      Appearance <- "VP 45"
   Polygon "Polygon_196" at 843,458 size 11x11
      Appearance <- "VP 45"
   Polygon "Polygon_199" at 630,469 size 11x11
      Appearance <- "VP 33"
   Polygon "Polygon_200" at 631,458 size 11x11
      Appearance <- "VP 33"
   Polygon "Polygon_157" at 417,469 size 11x11
      Appearance <- "VP 21"
   Polygon "Polygon_158" at 418,458 size 11x11
      Appearance <- "VP 21"
   Polygon "Polygon_151" at 205,469 size 11x11
      Appearance <- "VP 16"
   Polygon "Polygon_152" at 206,458 size 11x11
      Appearance <- "VP 16"
   Polygon "Polygon_201" at 83,465 size 11x11
      Appearance <- "VP 1"
   Polygon "Polygon_202" at 94,466 size 11x11
      Appearance <- "VP 1"
   Polygon "Polygon_5" at 83,508 size 11x11
      Appearance <- "VP 2"
   Polygon "Polygon_6" at 94,509 size 11x11
      Appearance <- "VP 2"
   Polygon "Polygon_7" at 83,551 size 11x11
      Appearance <- "VP 3"
   Polygon "Polygon_8" at 94,552 size 11x11
      Appearance <- "VP 3"
   Polygon "Polygon_9" at 83,595 size 11x11
      Appearance <- "VP 4"
   Polygon "Polygon_10" at 94,596 size 11x11
      Appearance <- "VP 4"
   Polygon "Polygon_11" at 124,490 size 11x11
      Appearance <- "VP 5"
   Polygon "Polygon_12" at 135,491 size 11x11
      Appearance <- "VP 5"
   Polygon "Polygon_13" at 158,490 size 11x11
      Appearance <- "VP 7"
   Polygon "Polygon_14" at 169,491 size 11x11
      Appearance <- "VP 7"
   Polygon "Polygon_15" at 124,576 size 11x11
      Appearance <- "VP 6"
   Polygon "Polygon_16" at 135,577 size 11x11
      Appearance <- "VP 6"
   Polygon "Polygon_207" at 158,576 size 11x11
      Appearance <- "VP 8"
   Polygon "Polygon_208" at 169,577 size 11x11
      Appearance <- "VP 8"
   Polygon "Polygon_17" at 295,465 size 11x11
      Appearance <- "VP 9"
   Polygon "Polygon_18" at 306,466 size 11x11
      Appearance <- "VP 9"
   Polygon "Polygon_19" at 295,508 size 11x11
      Appearance <- "VP 10"
   Polygon "Polygon_20" at 306,509 size 11x11
      Appearance <- "VP 10"
   Polygon "Polygon_21" at 295,551 size 11x11
      Appearance <- "VP 11"
   Polygon "Polygon_22" at 306,552 size 11x11
      Appearance <- "VP 11"
   Polygon "Polygon_23" at 295,595 size 11x11
      Appearance <- "VP 12"
   Polygon "Polygon_24" at 306,596 size 11x11
      Appearance <- "VP 12"
   Polygon "Polygon_25" at 336,490 size 11x11
      Appearance <- "VP 17"
   Polygon "Polygon_26" at 347,491 size 11x11
      Appearance <- "VP 17"
   Polygon "Polygon_27" at 370,490 size 11x11
      Appearance <- "VP 18"
   Polygon "Polygon_28" at 381,491 size 11x11
      Appearance <- "VP 18"
   Polygon "Polygon_29" at 336,576 size 11x11
      Appearance <- "VP 19"
   Polygon "Polygon_30" at 347,577 size 11x11
      Appearance <- "VP 19"
   Polygon "Polygon_31" at 370,576 size 11x11
      Appearance <- "VP 20"
   Polygon "Polygon_32" at 381,577 size 11x11
      Appearance <- "VP 20"
   Polygon "Polygon_33" at 507,465 size 11x11
      Appearance <- "VP 24"
   Polygon "Polygon_34" at 518,466 size 11x11
      Appearance <- "VP 24"
   Polygon "Polygon_35" at 507,508 size 11x11
      Appearance <- "VP 25"
   Polygon "Polygon_36" at 518,509 size 11x11
      Appearance <- "VP 25"
   Polygon "Polygon_37" at 507,551 size 11x11
      Appearance <- "VP 26"
   Polygon "Polygon_38" at 518,552 size 11x11
      Appearance <- "VP 26"
   Polygon "Polygon_39" at 507,595 size 11x11
      Appearance <- "VP 27"
   Polygon "Polygon_40" at 518,596 size 11x11
      Appearance <- "VP 27"
   Polygon "Polygon_41" at 548,490 size 11x11
      Appearance <- "VP 29"
   Polygon "Polygon_42" at 559,491 size 11x11
      Appearance <- "VP 29"
   Polygon "Polygon_43" at 582,490 size 11x11
      Appearance <- "VP 30"
   Polygon "Polygon_44" at 593,491 size 11x11
      Appearance <- "VP 30"
   Polygon "Polygon_45" at 548,576 size 11x11
      Appearance <- "VP 31"
   Polygon "Polygon_46" at 559,577 size 11x11
      Appearance <- "VP 31"
   Polygon "Polygon_47" at 582,576 size 11x11
      Appearance <- "VP 32"
   Polygon "Polygon_48" at 593,577 size 11x11
      Appearance <- "VP 32"
   Polygon "Polygon_49" at 719,465 size 11x11
      Appearance <- "VP 36"
   Polygon "Polygon_50" at 730,466 size 11x11
      Appearance <- "VP 36"
   Polygon "Polygon_51" at 719,508 size 11x11
      Appearance <- "VP 37"
   Polygon "Polygon_52" at 730,509 size 11x11
      Appearance <- "VP 37"
   Polygon "Polygon_53" at 719,551 size 11x11
      Appearance <- "VP 38"
   Polygon "Polygon_54" at 730,552 size 11x11
      Appearance <- "VP 38"
   Polygon "Polygon_55" at 719,595 size 11x11
      Appearance <- "VP 39"
   Polygon "Polygon_56" at 730,596 size 11x11
      Appearance <- "VP 39"
   Polygon "Polygon_57" at 760,490 size 11x11
      Appearance <- "VP 41"
   Polygon "Polygon_58" at 771,491 size 11x11
      Appearance <- "VP 41"
   Polygon "Polygon_59" at 794,490 size 11x11
      Appearance <- "VP 42"
   Polygon "Polygon_60" at 805,491 size 11x11
      Appearance <- "VP 42"
   Polygon "Polygon_61" at 760,576 size 11x11
      Appearance <- "VP 43"
   Polygon "Polygon_62" at 771,577 size 11x11
      Appearance <- "VP 43"
   Polygon "Polygon_63" at 794,576 size 11x11
      Appearance <- "VP 44"
   Polygon "Polygon_64" at 805,577 size 11x11
      Appearance <- "VP 44"
   Polygon "Polygon_65" at 931,465 size 11x11
      Appearance <- "VP 48"
   Polygon "Polygon_66" at 942,466 size 11x11
      Appearance <- "VP 48"
   Polygon "Polygon_67" at 931,508 size 11x11
      Appearance <- "VP 49"
   Polygon "Polygon_68" at 942,509 size 11x11
      Appearance <- "VP 49"
   Polygon "Polygon_69" at 931,551 size 11x11
      Appearance <- "VP 50"
   Polygon "Polygon_70" at 942,552 size 11x11
      Appearance <- "VP 50"
   Polygon "Polygon_71" at 931,595 size 11x11
      Appearance <- "VP 51"
   Polygon "Polygon_72" at 942,596 size 11x11
      Appearance <- "VP 51"
   Polygon "Polygon_73" at 972,490 size 11x11
      Appearance <- "VP 53"
   Polygon "Polygon_74" at 983,491 size 11x11
      Appearance <- "VP 53"
   Polygon "Polygon_75" at 1006,490 size 11x11
      Appearance <- "VP 54"
   Polygon "Polygon_76" at 1017,491 size 11x11
      Appearance <- "VP 54"
   Polygon "Polygon_77" at 972,576 size 11x11
      Appearance <- "VP 55"
   Polygon "Polygon_78" at 983,577 size 11x11
      Appearance <- "VP 55"
   Polygon "Polygon_79" at 1006,576 size 11x11
      Appearance <- "VP 56"
   Polygon "Polygon_80" at 1017,577 size 11x11
      Appearance <- "VP 56"
   Polygon "Polygon_81" at 1143,465 size 11x11
      Appearance <- "VP 60"
   Polygon "Polygon_82" at 1154,466 size 11x11
      Appearance <- "VP 60"
   Polygon "Polygon_83" at 1143,508 size 11x11
      Appearance <- "VP 61"
   Polygon "Polygon_84" at 1154,509 size 11x11
      Appearance <- "VP 61"
   Polygon "Polygon_85" at 1143,551 size 11x11
      Appearance <- "VP 62"
   Polygon "Polygon_86" at 1154,552 size 11x11
      Appearance <- "VP 62"
   Polygon "Polygon_87" at 1143,595 size 11x11
      Appearance <- "VP 63"
   Polygon "Polygon_88" at 1154,596 size 11x11
      Appearance <- "VP 63"
   Polygon "Polygon_89" at 1184,490 size 11x11
      Appearance <- "VP 65"
   Polygon "Polygon_90" at 1195,491 size 11x11
      Appearance <- "VP 65"
   Polygon "Polygon_91" at 1218,490 size 11x11
      Appearance <- "VP 66"
   Polygon "Polygon_92" at 1229,491 size 11x11
      Appearance <- "VP 66"
   Polygon "Polygon_93" at 1184,576 size 11x11
      Appearance <- "VP 67"
   Polygon "Polygon_94" at 1195,577 size 11x11
      Appearance <- "VP 67"
   Polygon "Polygon_95" at 1218,576 size 11x11
      Appearance <- "VP 68"
   Polygon "Polygon_96" at 1229,577 size 11x11
      Appearance <- "VP 68"
   Polygon "Polygon_97" at 1355,465 size 11x11
      Appearance <- "VP 72"
   Polygon "Polygon_98" at 1366,466 size 11x11
      Appearance <- "VP 72"
   Polygon "Polygon_99" at 1355,508 size 11x11
      Appearance <- "VP 73"
   Polygon "Polygon_100" at 1366,509 size 11x11
      Appearance <- "VP 73"
   Polygon "Polygon_101" at 1355,551 size 11x11
      Appearance <- "VP 74"
   Polygon "Polygon_102" at 1366,552 size 11x11
      Appearance <- "VP 74"
   Polygon "Polygon_103" at 1355,595 size 11x11
      Appearance <- "VP 75"
   Polygon "Polygon_104" at 1366,596 size 11x11
      Appearance <- "VP 75"
   Polygon "Polygon_105" at 1396,490 size 11x11
      Appearance <- "VP 77"
   Polygon "Polygon_106" at 1407,491 size 11x11
      Appearance <- "VP 77"
   Polygon "Polygon_107" at 1430,490 size 11x11
      Appearance <- "VP 78"
   Polygon "Polygon_108" at 1441,491 size 11x11
      Appearance <- "VP 78"
   Polygon "Polygon_109" at 1396,576 size 11x11
      Appearance <- "VP 79"
   Polygon "Polygon_110" at 1407,577 size 11x11
      Appearance <- "VP 79"
   Polygon "Polygon_111" at 1430,576 size 11x11
      Appearance <- "VP 80"
   Polygon "Polygon_112" at 1441,577 size 11x11
      Appearance <- "VP 80"
   Polygon "Polygon_113" at 142,942 size 11x11
      Appearance <- "VP 87"
   Polygon "Polygon_114" at 153,943 size 11x11
      Appearance <- "VP 87"
   Polygon "Polygon_3" at 30,890 size 11x11
      Appearance <- "VP 86"
   Polygon "Polygon_4" at 41,891 size 11x11
      Appearance <- "VP 86"
   Polygon "Polygon_115" at 123,352 size 58x419
      Visibility <- "step_vessel_1_proses"
      Appearance <- "VP 5"
   Line "Line_112" at 124,432 size 57x0
      Visibility <- "step_vessel_1_proses"
   Line "Line_113" at 142,385 size 21x0
      Visibility <- "step_vessel_1_proses"
   Line "Line_114" at 124,680 size 56x0
      Visibility <- "step_vessel_1_proses"
   Polygon "Polygon_116" at 335,352 size 58x419
      Appearance <- "VP 17"
      Visibility <- "step_vessel_2_proses"
   Line "Line_115" at 336,432 size 57x0
      Visibility <- "step_vessel_2_proses"
   Line "Line_116" at 354,385 size 21x0
      Visibility <- "step_vessel_2_proses"
   Line "Line_211" at 336,680 size 56x0
      Visibility <- "step_vessel_2_proses"
   Polygon "Polygon_189" at 547,352 size 58x419
      Appearance <- "VP 29"
      Visibility <- "step_vessel_3_proses"
   Line "Line_212" at 548,432 size 57x0
      Visibility <- "step_vessel_3_proses"
   Line "Line_213" at 566,385 size 21x0
      Visibility <- "step_vessel_3_proses"
   Line "Line_214" at 548,680 size 56x0
      Visibility <- "step_vessel_3_proses"
   Polygon "Polygon_190" at 759,352 size 58x419
      Appearance <- "VP 41"
      Visibility <- "step_vessel_4_proses"
   Line "Line_215" at 760,432 size 57x0
      Visibility <- "step_vessel_4_proses"
   Line "Line_216" at 778,385 size 21x0
      Visibility <- "step_vessel_4_proses"
   Line "Line_217" at 760,680 size 56x0
      Visibility <- "step_vessel_4_proses"
   Polygon "Polygon_203" at 971,352 size 58x419
      Appearance <- "VP 53"
      Visibility <- "step_vessel_5_proses"
   Line "Line_218" at 972,432 size 57x0
      Visibility <- "step_vessel_5_proses"
   Line "Line_219" at 990,385 size 21x0
      Visibility <- "step_vessel_5_proses"
   Line "Line_220" at 972,680 size 56x0
      Visibility <- "step_vessel_5_proses"
   Polygon "Polygon_204" at 1183,352 size 58x419
      Appearance <- "VP 65"
      Visibility <- "step_vessel_6_proses"
   Line "Line_221" at 1184,432 size 57x0
      Visibility <- "step_vessel_6_proses"
   Line "Line_222" at 1202,385 size 21x0
      Visibility <- "step_vessel_6_proses"
   Line "Line_223" at 1184,680 size 56x0
      Visibility <- "step_vessel_6_proses"
   Polygon "Polygon_209" at 1395,352 size 58x419
      Appearance <- "VP 77"
      Visibility <- "step_vessel_7_proses"
   Line "Line_224" at 1396,432 size 57x0
      Visibility <- "step_vessel_7_proses"
   Line "Line_225" at 1414,385 size 21x0
      Visibility <- "step_vessel_7_proses"
   Line "Line_226" at 1396,680 size 56x0
      Visibility <- "step_vessel_7_proses"
   IOField "I/O field_3" at 141,608 size 38x17; FormatPattern 9999999
   TextField "Text field_15" at 177,608 size 25x18; Text 'bar'
   IOField "I/O field_4" at 141,632 size 38x17; FormatPattern 9999999
   TextField "Text field_16" at 177,632 size 23x18; Text 'º C'
   IOField "I/O field_7" at 353,608 size 38x17; FormatPattern 9999999
   TextField "Text field_31" at 389,608 size 25x18; Text 'bar'
   IOField "I/O field_8" at 353,632 size 38x17; FormatPattern 9999999
   TextField "Text field_32" at 389,632 size 23x18; Text 'º C'
   IOField "I/O field_11" at 565,608 size 38x17; FormatPattern 9999999
   TextField "Text field_5" at 601,608 size 25x18; Text 'bar'
   IOField "I/O field_12" at 565,632 size 38x17; FormatPattern 9999999
   TextField "Text field_6" at 601,632 size 23x18; Text 'º C'
   IOField "I/O field_15" at 777,608 size 38x17; FormatPattern 9999999
   TextField "Text field_17" at 813,608 size 25x18; Text 'bar'
   IOField "I/O field_16" at 777,632 size 38x17; FormatPattern 9999999
   TextField "Text field_18" at 813,632 size 23x18; Text 'º C'
   IOField "I/O field_19" at 989,608 size 38x17; FormatPattern 9999999
   TextField "Text field_19" at 1025,608 size 25x18; Text 'bar'
   IOField "I/O field_20" at 989,632 size 38x17; FormatPattern 9999999
   TextField "Text field_20" at 1025,632 size 23x18; Text 'º C'
   IOField "I/O field_23" at 1201,608 size 38x17; FormatPattern 9999999
   TextField "Text field_21" at 1237,608 size 25x18; Text 'bar'
   IOField "I/O field_24" at 1201,632 size 38x17; FormatPattern 9999999
   TextField "Text field_22" at 1237,632 size 23x18; Text 'º C'
   IOField "I/O field_27" at 1413,608 size 38x17; FormatPattern 9999999
   TextField "Text field_23" at 1449,608 size 25x18; Text 'bar'
   IOField "I/O field_28" at 1413,632 size 38x17; FormatPattern 9999999
   TextField "Text field_24" at 1449,632 size 23x18; Text 'º C'
   Line "Line_1" at 109,467 size 0x141
      Appearance <- "step_vessel_1"
      Visibility <- "step_vessel_1_proses"
   Line "Line_3" at 110,496 size 16x0
      Appearance <- "step_vessel_1"
      Visibility <- "step_vessel_1_proses"
   Line "Line_4" at 110,582 size 16x0
      Appearance <- "step_vessel_1"
      Visibility <- "step_vessel_1_proses"
   Line "Line_17" at 321,466 size 0x157
      Appearance <- "step_vessel_2"
      Visibility <- "step_vessel_2_proses"
   Line "Line_18" at 318,496 size 16x0
      Appearance <- "step_vessel_2"
      Visibility <- "step_vessel_2_proses"
   Line "Line_19" at 318,582 size 16x0
      Appearance <- "step_vessel_2"
      Visibility <- "step_vessel_2_proses"
   Group "Tank vessel 1_1" at 123,352 size 58x419
   Group "Group_1" at 109,467 size 17x141
   Group "Group_76" at 180,475 size 118x150
   Group "Group_100" at 318,466 size 16x157
   Group "Tank vessel 2_1" at 335,352 size 58x419
   Group "Group_126" at 392,475 size 118x150
   Group "Group_148" at 605,475 size 118x150
   Group "Group_149" at 817,475 size 118x150
   Group "Group_150" at 1030,475 size 118x150
   Group "Group_151" at 1241,475 size 114x150
   Group "Group_152" at 1453,481 size 80x138
   Group "Group_86" at 739,620 size 12x22
   Group "Group_157" at 745,466 size 21x155
   Group "Group_155" at 533,466 size 17x154
   Group "Group_159" at 954,466 size 20x158
   Group "Group_161" at 1169,466 size 21x156
   Group "Group_163" at 1381,466 size 17x156
   Group "Group_5" at 536,400 size 40x99
   Group "Group_189" at 1172,400 size 40x99
   Polyline "Polyline_8" at 153,793 size 18x84
      Visibility <- "VB 1"
      Appearance <- "step_vessel_1_proses"
   Polyline "Polyline_11" at 365,793 size 18x84
      Visibility <- "VB 2"
      Appearance <- "step_vessel_2_proses"
   Polyline "Polyline_12" at 577,793 size 18x84
      Visibility <- "VB 3"
      Appearance <- "step_vessel_3_proses"
   Polyline "Polyline_14" at 789,793 size 18x84
      Visibility <- "VB 4"
      Appearance <- "step_vessel_4_proses"
   Polyline "Polyline_16" at 1001,793 size 18x84
      Visibility <- "VB 5"
      Appearance <- "step_vessel_5_proses"
   Polyline "Polyline_18" at 1213,793 size 18x84
      Visibility <- "VB 6"
      Appearance <- "step_vessel_6_proses"
   Polyline "Polyline_20" at 1425,793 size 18x84
      Visibility <- "VB 7"
      Appearance <- "step_vessel_7_proses"
   Group "Group_129" at 547,352 size 58x419
   Group "Group_144" at 759,352 size 58x419
   Group "Group_145" at 971,352 size 58x419
   Group "Group_146" at 1183,352 size 58x419
   Group "Group_147" at 1395,352 size 58x419
   Group "Tank vessel 1" at 123,352 size 58x419
   Group "Tank vessel 2" at 335,352 size 58x419
   Group "Group_116" at 547,352 size 58x419
   Group "Group_119" at 759,352 size 58x419
   Group "Group_120" at 971,352 size 58x419
   Group "Group_121" at 1183,352 size 58x419
   Group "Group_122" at 1395,352 size 58x419
   Group "Tank vessel 1_2" at 123,352 size 58x419
   Group "Tank vessel 2_2" at 335,352 size 58x419
   Group "Group_196" at 547,352 size 58x419
   Group "Group_197" at 759,352 size 58x419
   Group "Group_198" at 971,352 size 58x419
   Group "Group_200" at 1395,352 size 58x419
   Group "Group_199" at 1183,352 size 58x419
   Group "Group_127" at 420,640 size 1121x45
   Polygon "Polygon_210" at 123,352 size 58x419
      Visibility <- "step_vessel_1_proses"
      Appearance <- "step_vessel_1_proses"
   Line "Line_110" at 124,432 size 57x0
      Visibility <- "step_vessel_1_proses"
   Line "Line_111" at 142,385 size 21x0
      Visibility <- "step_vessel_1_proses"
   Line "Line_227" at 124,680 size 56x0
      Visibility <- "step_vessel_1_proses"
   Line "Line_228" at 112,400 size 25x11
      Visibility <- "VP 5"
      Appearance <- "step_vessel_1_proses"
   Line "Line_229" at 116,412 size 36x78
      Visibility <- "VP 5"
      Appearance <- "step_vessel_1_proses"
   Line "Line_230" at 152,488 size 0x11
      Visibility <- "VP 5"
      Appearance <- "step_vessel_1_proses"
   Line "Line_232" at 131,595 size 21x144
      Visibility <- "VP 5"
      Appearance <- "step_vessel_1_proses"
   Line "Line_233" at 152,579 size 0x19
      Visibility <- "VP 5"
      Appearance <- "step_vessel_1_proses"
   Line "Line_234" at 128,739 size 25x0
      Visibility <- "VP 5"
      Appearance <- "step_vessel_1_proses"
   Line "Line_236" at 105,898 size 0x48
      Visibility <- "step_vessel_1"
   Line "Line_237" at 102,948 size 40x0
      Visibility <- "step_vessel_1"
   Rectangle "Rectangle_3" at 75,874 size 1423x33
      Visibility <- "step_vessel_1"
   Line "Line_238" at 105,898 size 0x48
      Visibility <- "step_vessel_2"
   Line "Line_239" at 102,948 size 40x0
      Visibility <- "step_vessel_2"
   Rectangle "Rectangle_4" at 75,874 size 1423x33
      Visibility <- "step_vessel_2"
   Group "Preparation_out_2" at 75,874 size 1423x74
   Group "Preparation_out_1" at 75,874 size 1423x74
   Group "Preparation_out" at 75,874 size 1423x74
   Group "pipa_atas_vesel1_1" at 112,400 size 40x99
   Line "Line_231" at 146,496 size 12x0
      Visibility <- "VP 5"
      Appearance <- "step_vessel_1_proses"
   Line "Line_235" at 146,582 size 12x0
      Visibility <- "VP 5"
      Appearance <- "step_vessel_1_proses"
   Line "Line_270" at 358,582 size 12x0
      Visibility <- "step_vessel_2_proses"
      Appearance <- "step_vessel_2_proses"
   Line "Line_391" at 570,496 size 12x0
      Visibility <- "VP 29"
      Appearance <- "step_vessel_3_proses"
   Group "Group_176" at 536,400 size 40x99
   Line "Line_393" at 570,582 size 12x0
      Visibility <- "VP 29"
      Appearance <- "step_vessel_3_proses"
   Line "Line_204" at 782,582 size 12x0
      Visibility <- "VP 41"
      Appearance <- "step_vessel_4_proses"
   Line "Line_203" at 782,496 size 12x0
      Visibility <- "VP 41"
      Appearance <- "step_vessel_4_proses"
   Group "Group_7" at 748,400 size 40x99
   Line "Line_205" at 994,496 size 12x0
      Visibility <- "VP 53"
      Appearance <- "step_vessel_5_proses"
   Line "Line_206" at 994,582 size 12x0
      Visibility <- "VP 53"
      Appearance <- "step_vessel_5_proses"
   Line "Line_208" at 1206,582 size 15x0
      Visibility <- "VP 65"
      Appearance <- "step_vessel_6_proses"
   Line "Line_210" at 1418,582 size 12x0
      Visibility <- "VP 77"
      Appearance <- "step_vessel_7_proses"
   Line "Line_209" at 1418,496 size 12x0
      Visibility <- "VP 77"
      Appearance <- "step_vessel_7_proses"
   Group "Group_113" at 1384,400 size 40x99
   Group "Group_111" at 1172,400 size 40x99
   Line "Line_207" at 1206,496 size 17x0
      Visibility <- "VP 65"
      Appearance <- "step_vessel_6_proses"
   Line "Line_263" at 358,496 size 12x0
      Visibility <- "VP 17"
      Appearance <- "step_vessel_2_proses"
   Group "Group_109" at 960,400 size 40x99
   Group "Group_115" at 324,400 size 40x99
   Line "Line_240" at 105,898 size 0x48
      Visibility <- "step_vessel_3"
   Line "Line_241" at 102,948 size 40x0
      Visibility <- "step_vessel_3"
   Rectangle "Rectangle_5" at 75,874 size 1423x33
      Visibility <- "step_vessel_3"
   Group "Preparation_out_3" at 75,874 size 1423x74
   Group "pipa_atas_vesel1" at 112,400 size 40x99
   Line "Line_197" at 146,496 size 12x0
      Visibility <- "step_vessel_1_proses"
      Appearance <- "step_vessel_1"
   Line "Line_198" at 146,582 size 12x0
      Visibility <- "step_vessel_1_proses"
      Appearance <- "step_vessel_1"
   Line "Line_200" at 358,582 size 12x0
      Visibility <- "step_vessel_2_proses"
      Appearance <- "step_vessel_2"
   Line "Line_392" at 570,496 size 12x0
      Appearance <- "step_vessel_3"
      Visibility <- "step_vessel_3_proses"
   Group "Group_175" at 536,400 size 40x99
   Line "Line_394" at 570,582 size 12x0
      Appearance <- "step_vessel_3"
      Visibility <- "step_vessel_3_proses"
   Group "Group_182" at 960,400 size 40x99
   Line "Line_242" at 105,898 size 0x48
      Visibility <- "step_vessel_4"
   Line "Line_243" at 102,948 size 40x0
      Visibility <- "step_vessel_4"
   Rectangle "Rectangle_6" at 75,874 size 1423x33
      Visibility <- "step_vessel_4"
   Group "Preparation_out_4" at 75,874 size 1423x74
   Line "Line_244" at 105,898 size 0x48
      Visibility <- "step_vessel_5"
   Line "Line_245" at 102,948 size 40x0
      Visibility <- "step_vessel_5"
   Rectangle "Rectangle_7" at 75,874 size 1423x33
      Visibility <- "step_vessel_5"
   Group "Preparation_out_5" at 75,874 size 1423x74
   Group "Group_201" at 340,579 size 25x160
   Line "Line_246" at 105,898 size 0x48
      Visibility <- "step_vessel_6"
   Line "Line_247" at 102,948 size 40x0
      Visibility <- "step_vessel_6"
   Rectangle "Rectangle_8" at 75,874 size 1423x33
      Visibility <- "step_vessel_6"
   Group "Preparation_out_6" at 75,874 size 1423x74
   Group "Group_191" at 552,579 size 25x160
   Group "Group_192" at 764,579 size 25x160
   Group "Group_193" at 976,579 size 25x160
   Group "Group_195" at 1400,579 size 25x160
   Group "Group_194" at 1188,579 size 25x160
   Group "pipabawah_vessel1_1" at 128,579 size 25x160
   Group "Group_124" at 340,579 size 25x160
   Line "Line_248" at 105,898 size 0x48
      Visibility <- "step_vessel_7"
   Line "Line_249" at 102,948 size 40x0
      Visibility <- "step_vessel_7"
   Rectangle "Rectangle_9" at 75,874 size 1423x33
      Visibility <- "step_vessel_7"
   Line "Line_250" at 109,467 size 0x141
      Visibility <- "VP 5"
      Appearance <- "step_vessel_1_proses"
   Line "Line_251" at 110,496 size 16x0
      Visibility <- "VP 5"
      Appearance <- "step_vessel_1_proses"
   Line "Line_252" at 110,582 size 16x0
      Visibility <- "VP 5"
      Appearance <- "step_vessel_1_proses"
   Line "Line_253" at 180,582 size 30x0
      Visibility <- "VP 8"
   Line "Line_254" at 211,475 size 0x146
      Visibility <- "VP 8"
   Line "Line_255" at 213,600 size 85x0
      Visibility <- "VP 8"
   Line "Line_256" at 251,600 size 0x25
      Visibility <- "VP 8"
   Line "Line_257" at 321,466 size 0x157
      Appearance <- "step_vessel_2_proses"
      Visibility <- "VP 17"
   Line "Line_258" at 318,496 size 16x0
      Appearance <- "step_vessel_2_proses"
      Visibility <- "VP 17"
   Line "Line_259" at 318,582 size 16x0
      Appearance <- "step_vessel_2_proses"
      Visibility <- "VP 17"
   Polygon "Polygon_211" at 335,352 size 58x419
      Appearance <- "step_vessel_2_proses"
      Visibility <- "step_vessel_2_proses"
   Line "Line_260" at 336,432 size 57x0
      Visibility <- "step_vessel_2_proses"
   Line "Line_261" at 354,385 size 21x0
      Visibility <- "step_vessel_2_proses"
   Line "Line_262" at 336,680 size 56x0
      Visibility <- "step_vessel_2_proses"
   Line "Line_264" at 324,400 size 25x11
      Visibility <- "VP 17"
      Appearance <- "step_vessel_2_proses"
   Line "Line_265" at 328,412 size 36x78
      Visibility <- "VP 17"
      Appearance <- "step_vessel_2_proses"
   Line "Line_266" at 364,488 size 0x11
      Visibility <- "VP 17"
      Appearance <- "step_vessel_2_proses"
   Line "Line_267" at 343,595 size 21x144
      Appearance <- "step_vessel_2_proses"
      Visibility <- "VP 17"
   Line "Line_268" at 364,579 size 0x19
      Appearance <- "step_vessel_2_proses"
      Visibility <- "VP 17"
   Line "Line_269" at 340,739 size 25x0
      Appearance <- "step_vessel_2_proses"
      Visibility <- "VP 17"
   Group "Group_128" at 420,640 size 1121x45
   Line "Line_276" at 1538,684 size 0x259
      Visibility <- "VP 22"
   Line "Line_274" at 423,640 size 0x45
      Visibility <- "VP 22"
   Line "Line_275" at 420,683 size 1121x0
      Visibility <- "VP 22"
   Polygon "Polygon_212" at 547,352 size 58x419
      Appearance <- "step_vessel_3_proses"
      Visibility <- "step_vessel_3_proses"
   Line "Line_277" at 548,432 size 57x0
      Visibility <- "step_vessel_3_proses"
   Line "Line_278" at 566,385 size 21x0
      Visibility <- "step_vessel_3_proses"
   Line "Line_279" at 548,680 size 56x0
      Visibility <- "step_vessel_3_proses"
   Line "Line_280" at 636,643 size 0x42
      Visibility <- "VP 34"
   Line "Line_281" at 634,683 size 907x0
      Visibility <- "VP 34"
   Line "Line_282" at 1538,680 size 0x261
      Visibility <- "VP 34"
   Group "Group_138" at 634,643 size 907x298
   Group "Group_140" at 845,643 size 695x299
   Group "Group_141" at 1058,642 size 483x294
   Group "Group_142" at 1272,642 size 269x301
   Group "Group_143" at 1484,643 size 56x300
   Group "Group_133" at 777,608 size 61x42
   Group "Group_172" at 208,643 size 1333x301
   Group "Group_139" at 420,640 size 1121x303
   Group "Group_78" at 417,620 size 12x22
   Group "proses_2" at 75,874 size 1423x74
   Line "Line_283" at 848,643 size 0x38
      Visibility <- "VP 46"
   Line "Line_284" at 845,683 size 695x0
      Visibility <- "VP 46"
   Line "Line_285" at 1538,680 size 0x262
      Visibility <- "VP 46"
   Line "Line_286" at 1061,642 size 0x44
      Visibility <- "VP 58"
   Line "Line_287" at 1058,683 size 483x0
      Visibility <- "VP 58"
   Line "Line_288" at 1538,681 size 0x255
      Visibility <- "VP 58"
   Line "Line_291" at 1538,680 size 0x263
      Visibility <- "VP 70"
   Line "Line_290" at 1272,683 size 269x0
      Visibility <- "VP 70"
   Line "Line_289" at 1275,642 size 0x38
      Visibility <- "VP 70"
   Line "Line_292" at 1487,643 size 0x38
      Visibility <- "VP 82"
   Line "Line_294" at 1484,683 size 56x0
      Visibility <- "VP 82"
   Line "Line_293" at 1538,680 size 0x263
      Visibility <- "VP 82"
   Polygon "Polygon_213" at 759,352 size 58x419
      Appearance <- "step_vessel_4_proses"
      Visibility <- "step_vessel_4_proses"
   Line "Line_295" at 760,432 size 57x0
      Visibility <- "step_vessel_4_proses"
   Line "Line_296" at 778,385 size 21x0
      Visibility <- "step_vessel_4_proses"
   Line "Line_297" at 760,680 size 56x0
      Visibility <- "step_vessel_4_proses"
   Polygon "Polygon_214" at 971,352 size 58x419
      Appearance <- "step_vessel_5_proses"
      Visibility <- "step_vessel_5_proses"
   Line "Line_117" at 972,432 size 57x0
      Visibility <- "step_vessel_5_proses"
   Line "Line_298" at 990,385 size 21x0
      Visibility <- "step_vessel_5_proses"
   Line "Line_299" at 972,680 size 56x0
      Visibility <- "step_vessel_5_proses"
   Polygon "Polygon_215" at 1183,352 size 58x419
      Appearance <- "step_vessel_6_proses"
      Visibility <- "step_vessel_6_proses"
   Line "Line_300" at 1184,432 size 57x0
      Visibility <- "step_vessel_6_proses"
   Line "Line_301" at 1202,385 size 21x0
      Visibility <- "step_vessel_6_proses"
   Line "Line_302" at 1184,680 size 56x0
      Visibility <- "step_vessel_6_proses"
   Polygon "Polygon_216" at 1395,352 size 58x419
      Appearance <- "step_vessel_7_proses"
      Visibility <- "step_vessel_7_proses"
   Line "Line_303" at 1396,432 size 57x0
      Visibility <- "step_vessel_7_proses"
   Line "Line_304" at 1414,385 size 21x0
      Visibility <- "step_vessel_7_proses"
   Line "Line_305" at 1396,680 size 56x0
      Visibility <- "step_vessel_7_proses"
   Line "Line_272" at 392,582 size 30x0
      Visibility <- "VP 20"
   Line "Line_273" at 423,475 size 0x146
      Visibility <- "VP 20"
   Line "Line_306" at 425,600 size 85x0
      Visibility <- "VP 20"
   Line "Line_307" at 463,600 size 0x25
      Visibility <- "VP 20"
   Line "Line_308" at 605,582 size 30x0
      Visibility <- "VP 32"
   Line "Line_309" at 636,475 size 0x146
      Visibility <- "VP 32"
   Line "Line_310" at 638,600 size 85x0
      Visibility <- "VP 32"
   Line "Line_311" at 676,600 size 0x25
      Visibility <- "VP 32"
   Line "Line_312" at 817,582 size 30x0
      Visibility <- "VP 44"
   Line "Line_313" at 848,475 size 0x146
      Visibility <- "VP 44"
   Line "Line_314" at 850,600 size 85x0
      Visibility <- "VP 44"
   Line "Line_315" at 888,600 size 0x25
      Visibility <- "VP 44"
   Line "Line_316" at 1030,582 size 30x0
      Visibility <- "VP 56"
   Line "Line_317" at 1061,475 size 0x146
      Visibility <- "VP 56"
   Line "Line_318" at 1063,600 size 85x0
      Visibility <- "VP 56"
   Line "Line_319" at 1099,600 size 0x25
      Visibility <- "VP 56"
   Line "Line_320" at 1241,582 size 33x0
      Visibility <- "VP 68"
   Line "Line_321" at 1275,475 size 0x146
      Visibility <- "VP 68"
   Line "Line_322" at 1277,600 size 78x0
      Visibility <- "VP 68"
   Line "Line_323" at 1311,600 size 0x25
      Visibility <- "VP 68"
   Line "Line_324" at 1453,582 size 33x0
      Visibility <- "VP 80"
   Line "Line_325" at 1487,481 size 0x138
      Visibility <- "VP 80"
   Line "Line_326" at 1489,600 size 44x0
      Visibility <- "VP 80"
   Line "Line_327" at 1524,600 size 0x19
      Visibility <- "VP 80"
   Line "Line_329" at 321,466 size 0x154
      Visibility <- "VP 17"
   Line "Line_330" at 318,496 size 16x0
      Visibility <- "VP 17"
   Line "Line_331" at 318,582 size 16x0
      Visibility <- "VP 17"
   Line "Line_332" at 533,466 size 0x154
      Visibility <- "VP 29"
      Appearance <- "step_vessel_3_proses"
   Line "Line_333" at 534,496 size 16x0
      Visibility <- "VP 29"
      Appearance <- "step_vessel_3_proses"
   Line "Line_334" at 534,582 size 16x0
      Visibility <- "VP 29"
      Appearance <- "step_vessel_3_proses"
   Group "Group_156" at 745,466 size 21x155
   Group "Group_154" at 533,466 size 17x157
   Group "Group_158" at 954,466 size 20x158
   Group "Group_160" at 1169,466 size 21x156
   Group "Group_162" at 1381,466 size 17x156
   Group "Group_137" at 109,467 size 17x141
   Group "Group_123" at 318,466 size 16x157
   Polyline "Polyline_1" at 153,793 size 18x84
      Appearance <- "VB 1"
      Visibility <- "step_vessel_1_proses"
   Polyline "Polyline_10" at 365,793 size 18x84
      Appearance <- "VB 2"
      Visibility <- "step_vessel_2_proses"
   Polyline "Polyline_13" at 577,793 size 18x84
      Appearance <- "VB 3"
      Visibility <- "step_vessel_3_proses"
   Polyline "Polyline_15" at 789,793 size 18x84
      Appearance <- "VB 4"
      Visibility <- "step_vessel_4_proses"
   Polyline "Polyline_17" at 1001,793 size 18x84
      Appearance <- "VB 5"
      Visibility <- "step_vessel_5_proses"
   Polyline "Polyline_19" at 1213,793 size 18x84
      Appearance <- "VB 6"
      Visibility <- "step_vessel_6_proses"
   Polyline "Polyline_21" at 1425,793 size 18x84
      Appearance <- "VB 7"
      Visibility <- "step_vessel_7_proses"
   Group "Group_187" at 748,400 size 40x99
   Line "Line_448" at 570,496 size 12x0
      Appearance <- "step_vessel_3"
   Line "Line_449" at 570,582 size 12x0
      Appearance <- "step_vessel_3"
   Group "Group_186" at 536,400 size 40x99
   Line "Line_447" at 782,496 size 12x0
      Appearance <- "step_vessel_4"
   Line "Line_456" at 782,582 size 12x0
      Appearance <- "step_vessel_4"
   Group "Group_188" at 960,400 size 40x99
   Group "pipa_atas_vesel1_2" at 112,400 size 40x99
   Line "Line_371" at 146,496 size 12x0
      Appearance <- "step_vessel_1"
   Group "pipabawah_vesel_2" at 128,579 size 25x160
   Line "Line_446" at 994,496 size 12x0
      Appearance <- "step_vessel_5"
   Line "Line_503" at 994,582 size 12x0
      Appearance <- "step_vessel_5"
   Line "Line_460" at 1206,582 size 15x0
      Appearance <- "step_vessel_6"
   Line "Line_467" at 1418,582 size 12x0
      Appearance <- "step_vessel_7"
   Line "Line_444" at 1418,496 size 12x0
      Appearance <- "step_vessel_7"
   Group "Group_190" at 1384,400 size 40x99
   Line "Line_445" at 1206,496 size 17x0
      Appearance <- "step_vessel_6"
   Line "Line_201" at 570,496 size 12x0
      Appearance <- "step_vessel_3"
   Group "Group_173" at 324,400 size 40x99
   Line "Line_504" at 358,496 size 12x0
      Appearance <- "step_vessel_2"
   Group "Group_174" at 1172,400 size 40x99
   Line "Line_335" at 745,466 size 0x155
      Visibility <- "VP 41"
      Appearance <- "step_vessel_4_proses"
   Line "Line_336" at 746,582 size 20x0
      Visibility <- "VP 41"
      Appearance <- "step_vessel_4_proses"
   Line "Line_337" at 747,496 size 19x0
      Visibility <- "VP 41"
      Appearance <- "step_vessel_4_proses"
   Line "Line_338" at 957,466 size 0x158
      Visibility <- "VP 53"
      Appearance <- "step_vessel_5_proses"
   Line "Line_339" at 955,496 size 19x0
      Visibility <- "VP 53"
      Appearance <- "step_vessel_5_proses"
   Line "Line_340" at 954,582 size 20x0
      Visibility <- "VP 53"
      Appearance <- "step_vessel_5_proses"
   Line "Line_341" at 1169,466 size 0x156
      Appearance <- "step_vessel_6_proses"
      Visibility <- "VP 65"
   Line "Line_342" at 1169,496 size 21x0
      Appearance <- "step_vessel_6_proses"
      Visibility <- "VP 65"
   Line "Line_343" at 1171,582 size 19x0
      Appearance <- "step_vessel_6_proses"
      Visibility <- "VP 65"
   Line "Line_344" at 1381,466 size 0x156
      Appearance <- "step_vessel_7_proses"
      Visibility <- "VP 77"
   Line "Line_345" at 1382,496 size 16x0
      Appearance <- "step_vessel_7_proses"
      Visibility <- "VP 77"
   Line "Line_346" at 1383,582 size 14x0
      Appearance <- "step_vessel_7_proses"
      Visibility <- "VP 77"
   Line "Line_347" at 745,466 size 0x155
      Appearance <- "step_vessel_4"
   Line "Line_348" at 746,582 size 20x0
      Appearance <- "step_vessel_4"
   Line "Line_349" at 747,496 size 19x0
      Appearance <- "step_vessel_4"
   Line "Line_350" at 533,466 size 0x157
      Appearance <- "step_vessel_3"
   Line "Line_351" at 534,496 size 16x0
      Appearance <- "step_vessel_3"
   Line "Line_352" at 534,582 size 16x0
      Appearance <- "step_vessel_3"
   Line "Line_353" at 957,466 size 0x158
      Appearance <- "step_vessel_5"
   Line "Line_354" at 955,496 size 19x0
      Appearance <- "step_vessel_5"
   Line "Line_355" at 954,582 size 20x0
      Appearance <- "step_vessel_5"
   Line "Line_356" at 1169,466 size 0x156
      Appearance <- "step_vessel_6"
   Line "Line_357" at 1169,496 size 21x0
      Appearance <- "step_vessel_6"
   Line "Line_358" at 1171,582 size 19x0
      Appearance <- "step_vessel_6"
   Line "Line_359" at 1381,466 size 0x156
      Appearance <- "step_vessel_7"
   Line "Line_360" at 1382,496 size 16x0
      Appearance <- "step_vessel_7"
   Line "Line_361" at 1383,582 size 14x0
      Appearance <- "step_vessel_7"
   Line "Line_362" at 109,467 size 0x141
      Appearance <- "step_vessel_1"
   Line "Line_363" at 110,496 size 16x0
      Appearance <- "step_vessel_1"
   Line "Line_364" at 110,582 size 16x0
      Appearance <- "step_vessel_1"
   Line "Line_365" at 321,466 size 0x157
      Appearance <- "step_vessel_2"
   Line "Line_366" at 318,496 size 16x0
      Appearance <- "step_vessel_2"
   Line "Line_367" at 318,582 size 16x0
      Appearance <- "step_vessel_2"
   Line "Line_368" at 112,400 size 25x11
      Appearance <- "step_vessel_1"
   Line "Line_369" at 116,412 size 36x78
      Appearance <- "step_vessel_1"
   Line "Line_370" at 152,488 size 0x11
      Appearance <- "step_vessel_1"
   Line "Line_372" at 131,595 size 21x144
      Appearance <- "step_vessel_1"
   Line "Line_373" at 152,579 size 0x19
      Appearance <- "step_vessel_1"
   Line "Line_374" at 128,739 size 25x0
      Appearance <- "step_vessel_1"
   Line "Line_378" at 1538,680 size 0x264
      Visibility <- "VP 13"
   Line "Line_377" at 208,683 size 1333x0
      Visibility <- "VP 13"
   Line "Line_376" at 211,643 size 0x38
      Visibility <- "VP 13"
   Line "Line_382" at 1172,400 size 25x11
      Appearance <- "step_vessel_6"
   Line "Line_383" at 1176,412 size 36x78
      Appearance <- "step_vessel_6"
   Line "Line_384" at 1212,488 size 0x11
      Appearance <- "step_vessel_6"
   Line "Line_385" at 536,400 size 25x11
      Appearance <- "step_vessel_3"
      Visibility <- "step_vessel_3_proses"
   Line "Line_386" at 540,412 size 36x78
      Appearance <- "step_vessel_3"
      Visibility <- "step_vessel_3_proses"
   Line "Line_387" at 576,488 size 0x11
      Appearance <- "step_vessel_3"
      Visibility <- "step_vessel_3_proses"
   Line "Line_388" at 536,400 size 25x11
      Visibility <- "VP 29"
      Appearance <- "step_vessel_3_proses"
   Line "Line_389" at 540,412 size 36x78
      Visibility <- "VP 29"
      Appearance <- "step_vessel_3_proses"
   Line "Line_390" at 576,488 size 0x11
      Visibility <- "VP 29"
      Appearance <- "step_vessel_3_proses"
   Line "Line_202" at 555,595 size 21x144
      Appearance <- "step_vessel_3"
      Visibility <- "step_vessel_3_proses"
   Line "Line_395" at 576,579 size 0x19
      Appearance <- "step_vessel_3"
      Visibility <- "step_vessel_3_proses"
   Line "Line_396" at 552,739 size 25x0
      Appearance <- "step_vessel_3"
      Visibility <- "step_vessel_3_proses"
   Line "Line_397" at 1384,400 size 25x11
      Appearance <- "step_vessel_7"
      Visibility <- "step_vessel_7_proses"
   Line "Line_398" at 1388,412 size 36x78
      Appearance <- "step_vessel_7"
      Visibility <- "step_vessel_7_proses"
   Line "Line_399" at 1424,488 size 0x11
      Appearance <- "step_vessel_7"
      Visibility <- "step_vessel_7_proses"
   Line "Line_401" at 1403,595 size 21x144
      Appearance <- "step_vessel_7"
      Visibility <- "step_vessel_7_proses"
   Line "Line_402" at 1424,579 size 0x19
      Appearance <- "step_vessel_7"
      Visibility <- "step_vessel_7_proses"
   Line "Line_403" at 1400,739 size 25x0
      Appearance <- "step_vessel_7"
      Visibility <- "step_vessel_7_proses"
   Line "Line_406" at 1191,595 size 21x144
      Appearance <- "step_vessel_6"
      Visibility <- "step_vessel_6_proses"
   Line "Line_407" at 1212,579 size 0x19
      Appearance <- "step_vessel_6"
      Visibility <- "step_vessel_6_proses"
   Line "Line_408" at 1188,739 size 25x0
      Appearance <- "step_vessel_6"
      Visibility <- "step_vessel_6_proses"
   Line "Line_410" at 1172,400 size 25x11
      Visibility <- "step_vessel_6_proses"
      Appearance <- "step_vessel_6"
   Line "Line_411" at 1176,412 size 36x78
      Appearance <- "step_vessel_6"
      Visibility <- "step_vessel_6_proses"
   Line "Line_412" at 1212,488 size 0x11
      Appearance <- "step_vessel_6"
      Visibility <- "step_vessel_6_proses"
   Line "Line_414" at 960,400 size 25x11
      Appearance <- "step_vessel_5"
      Visibility <- "step_vessel_5_proses"
   Line "Line_415" at 964,412 size 36x78
      Appearance <- "step_vessel_5"
      Visibility <- "step_vessel_5_proses"
   Line "Line_416" at 1000,488 size 0x11
      Appearance <- "step_vessel_5"
      Visibility <- "step_vessel_5_proses"
   Line "Line_418" at 979,595 size 21x144
      Appearance <- "step_vessel_5"
      Visibility <- "step_vessel_5_proses"
   Line "Line_419" at 1000,579 size 0x19
      Appearance <- "step_vessel_5"
      Visibility <- "step_vessel_5_proses"
